// TIA Portal project "XSFW_TIA60401_A2" (V13) (continued)
VERSION : 0.1
   VAR
      x : Bool;
      x1 : Bool;
      x2 : Bool;
      x3 : Bool;
      x4 : Bool;
      x5 : Bool;
      x6 : Bool;
      x7 : Bool;
      x8 : Bool;
      x9 : Bool;
      x10 : Bool;
      x11 : Bool;
      x12 : Bool;
      x13 : Bool;
      x14 : Bool;
      x15 : Bool;
      x16 : Bool;
      x17 : Bool;
      x18 : Bool;
      x19 : Bool;
      x20 : Bool;
      x21 : Bool;
      x22 : Bool;
      x23 : Bool;
      x24 : Bool;
      x25 : Bool;
      x26 : Bool;
      x27 : Bool;
      x28 : Bool;
      x29 : Bool;
      x30 : Bool;
      x31 : Bool;
      x32 : Bool;
      x33 : Bool;
      x34 : Bool;
      x35 : Bool;
      x36 : Bool;
      x37 : Bool;
      x38 : Bool;
      x39 : Bool;
      x40 : Bool;
      x41 : Bool;
      x42 : Bool;
      x43 : Bool;
      x44 : Bool;
      x45 : Bool;
      x46 : Bool;
      x47 : Bool;
      x48 : Bool;
      x49 : Bool;
      x50 : Bool;
      x51 : Bool;
      x52 : Bool;
      x53 : Bool;
      x54 : Bool;
      x55 : Bool;
      x56 : Bool;
      x57 : Bool;
      x58 : Bool;
      x59 : Bool;
      x60 : Bool;
      x61 : Bool;
      x62 : Bool;
      x63 : Bool;
      x64 : Bool;
      x65 : Bool;
      x66 : Bool;
      x67 : Bool;
      x68 : Bool;
      x69 : Bool;
      x70 : Bool;
      x71 : Bool;
      x72 : Bool;
      x73 : Bool;
      x74 : Bool;
      x75 : Bool;
      x76 : Bool;
      x77 : Bool;
      x78 : Bool;
      x79 : Bool;
      x80 : Bool;
      x81 : Bool;
      x82 : Bool;
      x83 : Bool;
      x84 : Bool;
      x85 : Bool;
      x86 : Bool;
      x87 : Bool;
      x88 : Bool;
      x89 : Bool;
      x90 : Bool;
      x91 : Bool;
      x92 : Bool;
      x93 : Bool;
      x94 : Bool;
      x95 : Bool;
      x96 : Bool;
      x97 : Bool;
      x98 : Bool;
      x99 : Bool;
      x100 : Bool;
      x101 : Bool;
      x102 : Bool;
      x103 : Bool;
      x104 : Bool;
      x105 : Bool;
      x106 : Bool;
      x107 : Bool;
      x108 : Bool;
      x109 : Bool;
      x110 : Bool;
      x111 : Bool;
      x112 : Bool;
      x113 : Bool;
      x114 : Bool;
      x115 : Bool;
      x116 : Bool;
      x117 : Bool;
      x118 : Bool;
      x119 : Bool;
      x120 : Bool;
      x121 : Bool;
      x122 : Bool;
      x123 : Bool;
      x124 : Bool;
      x125 : Bool;
      x126 : Bool;
      x127 : Bool;
      x128 : Bool;
      x129 : Bool;
      x130 : Bool;
      x131 : Bool;
      x132 : Bool;
      x133 : Bool;
      x134 : Bool;
      x135 : Bool;
      x136 : Bool;
      x137 : Bool;
      x138 : Bool;
      x139 : Bool;
      x140 : Bool;
      x141 : Bool;
      x142 : Bool;
      x143 : Bool;
      x144 : Bool;
      x145 : Bool;
      x146 : Bool;
      x147 : Bool;
      x148 : Bool;
      x149 : Bool;
      x150 : Bool;
      x151 : Bool;
      x152 : Bool;
      x153 : Bool;
      x154 : Bool;
      x155 : Bool;
      x156 : Bool;
      x157 : Bool;
      x158 : Bool;
      x159 : Bool;
      x160 : Bool;
      x161 : Bool;
      x162 : Bool;
      x163 : Bool;
      x164 : Bool;
      x165 : Bool;
      x166 : Bool;
      x167 : Bool;
      x168 : Bool;
      x169 : Bool;
      x170 : Bool;
      x171 : Bool;
      x172 : Bool;
      x173 : Bool;
      x174 : Bool;
      x175 : Bool;
      x176 : Bool;
      x177 : Bool;
      x178 : Bool;
      x179 : Bool;
      x180 : Bool;
      x181 : Bool;
      x182 : Bool;
      x183 : Bool;
      x184 : Bool;
      x185 : Bool;
      x186 : Bool;
      x187 : Bool;
      x188 : Bool;
      x189 : Bool;
      x190 : Bool;
      x191 : Bool;
      x192 : Bool;
      x193 : Bool;
      x194 : Bool;
      x195 : Bool;
      x196 : Bool;
      x197 : Bool;
      x198 : Bool;
      x199 : Bool;
   END_VAR
BEGIN
END_DATA_BLOCK

DATA_BLOCK "DB_COM_REC_AUX"   // DB37
{ S7_Optimized_Access := 'FALSE' }
VERSION : 0.1
   VAR
      x : Bool;
      x1 : Bool;
      x2 : Bool;
      x3 : Bool;
      x4 : Bool;
      x5 : Bool;
      x6 : Bool;
      x7 : Bool;
      x8 : Bool;
      x9 : Bool;
      x10 : Bool;
      x11 : Bool;
      x12 : Bool;
      x13 : Bool;
      x14 : Bool;
      x15 : Bool;
      x16 : Bool;
      x17 : Bool;
      x18 : Bool;
      x19 : Bool;
      x20 : Bool;
      x21 : Bool;
      x22 : Bool;
      x23 : Bool;
      x24 : Bool;
      x25 : Bool;
      x26 : Bool;
      x27 : Bool;
      x28 : Bool;
      x29 : Bool;
      x30 : Bool;
      x31 : Bool;
      x32 : Bool;
      x33 : Bool;
      x34 : Bool;
      x35 : Bool;
      x36 : Bool;
      x37 : Bool;
      x38 : Bool;
      x39 : Bool;
      x40 : Bool;
      x41 : Bool;
      x42 : Bool;
      x43 : Bool;
      x44 : Bool;
      x45 : Bool;
      x46 : Bool;
      x47 : Bool;
      x48 : Bool;
      x49 : Bool;
      x50 : Bool;
      x51 : Bool;
      x52 : Bool;
      x53 : Bool;
      x54 : Bool;
      x55 : Bool;
      x56 : Bool;
      x57 : Bool;
      x58 : Bool;
      x59 : Bool;
      x60 : Bool;
      x61 : Bool;
      x62 : Bool;
      x63 : Bool;
      x64 : Bool;
      x65 : Bool;
      x66 : Bool;
      x67 : Bool;
      x68 : Bool;
      x69 : Bool;
      x70 : Bool;
      x71 : Bool;
      x72 : Bool;
      x73 : Bool;
      x74 : Bool;
      x75 : Bool;
      x76 : Bool;
      x77 : Bool;
      x78 : Bool;
      x79 : Bool;
      x80 : Bool;
      x81 : Bool;
      x82 : Bool;
      x83 : Bool;
      x84 : Bool;
      x85 : Bool;
      x86 : Bool;
      x87 : Bool;
      x88 : Bool;
      x89 : Bool;
      x90 : Bool;
      x91 : Bool;
      x92 : Bool;
      x93 : Bool;
      x94 : Bool;
      x95 : Bool;
      x96 : Bool;
      x97 : Bool;
      x98 : Bool;
      x99 : Bool;
      x100 : Bool;
      x101 : Bool;
      x102 : Bool;
      x103 : Bool;
      x104 : Bool;
      x105 : Bool;
      x106 : Bool;
      x107 : Bool;
      x108 : Bool;
      x109 : Bool;
      x110 : Bool;
      x111 : Bool;
      x112 : Bool;
      x113 : Bool;
      x114 : Bool;
      x115 : Bool;
      x116 : Bool;
      x117 : Bool;
      x118 : Bool;
      x119 : Bool;
      x120 : Bool;
      x121 : Bool;
      x122 : Bool;
      x123 : Bool;
      x124 : Bool;
      x125 : Bool;
      x126 : Bool;
      x127 : Bool;
      x128 : Bool;
      x129 : Bool;
      x130 : Bool;
      x131 : Bool;
      x132 : Bool;
      x133 : Bool;
      x134 : Bool;
      x135 : Bool;
      x136 : Bool;
      x137 : Bool;
      x138 : Bool;
      x139 : Bool;
      x140 : Bool;
      x141 : Bool;
      x142 : Bool;
      x143 : Bool;
      x144 : Bool;
      x145 : Bool;
      x146 : Bool;
      x147 : Bool;
      x148 : Bool;
      x149 : Bool;
      x150 : Bool;
      x151 : Bool;
      x152 : Bool;
      x153 : Bool;
      x154 : Bool;
      x155 : Bool;
      x156 : Bool;
      x157 : Bool;
      x158 : Bool;
      x159 : Bool;
      x160 : Bool;
      x161 : Bool;
      x162 : Bool;
      x163 : Bool;
      x164 : Bool;
      x165 : Bool;
      x166 : Bool;
      x167 : Bool;
      x168 : Bool;
      x169 : Bool;
      x170 : Bool;
      x171 : Bool;
      x172 : Bool;
      x173 : Bool;
      x174 : Bool;
      x175 : Bool;
      x176 : Bool;
      x177 : Bool;
      x178 : Bool;
      x179 : Bool;
      x180 : Bool;
      x181 : Bool;
      x182 : Bool;
      x183 : Bool;
      x184 : Bool;
      x185 : Bool;
      x186 : Bool;
      x187 : Bool;
      x188 : Bool;
      x189 : Bool;
      x190 : Bool;
      x191 : Bool;
      x192 : Bool;
      x193 : Bool;
      x194 : Bool;
      x195 : Bool;
      x196 : Bool;
      x197 : Bool;
      x198 : Bool;
      x199 : Bool;
   END_VAR
BEGIN
END_DATA_BLOCK

DATA_BLOCK "DB_BIT_VIDA"   // DB38
{ S7_Optimized_Access := 'FALSE' }
VERSION : 0.1
   VAR
      x : Bool;
      x1 : Bool;
      x2 : Bool;
      x3 : Bool;
      x4 : Bool;
      x5 : Bool;
      x6 : Bool;
      x7 : Bool;
      x8 : Bool;
      x9 : Bool;
      x10 : Bool;
      x11 : Bool;
      x12 : Bool;
      x13 : Bool;
      x14 : Bool;
      x15 : Bool;
      x16 : Bool;
      x17 : Bool;
      x18 : Bool;
      x19 : Bool;
      x20 : Bool;
      x21 : Bool;
      x22 : Bool;
      x23 : Bool;
      x24 : Bool;
      x25 : Bool;
      x26 : Bool;
      x27 : Bool;
      x28 : Bool;
      x29 : Bool;
      x30 : Bool;
      x31 : Bool;
      x32 : Bool;
      x33 : Bool;
      x34 : Bool;
      x35 : Bool;
      x36 : Bool;
      x37 : Bool;
      x38 : Bool;
      x39 : Bool;
      x40 : Bool;
      x41 : Bool;
      x42 : Bool;
      x43 : Bool;
      x44 : Bool;
      x45 : Bool;
      x46 : Bool;
      x47 : Bool;
      x48 : Bool;
      x49 : Bool;
      x50 : Bool;
      x51 : Bool;
      x52 : Bool;
      x53 : Bool;
      x54 : Bool;
      x55 : Bool;
      x56 : Bool;
      x57 : Bool;
      x58 : Bool;
      x59 : Bool;
      x60 : Bool;
      x61 : Bool;
      x62 : Bool;
      x63 : Bool;
      x64 : Bool;
      x65 : Bool;
      x66 : Bool;
      x67 : Bool;
      x68 : Bool;
      x69 : Bool;
      x70 : Bool;
      x71 : Bool;
      x72 : Bool;
      x73 : Bool;
      x74 : Bool;
      x75 : Bool;
      x76 : Bool;
      x77 : Bool;
      x78 : Bool;
      x79 : Bool;
      x80 : Bool;
      x81 : Bool;
      x82 : Bool;
      x83 : Bool;
      x84 : Bool;
      x85 : Bool;
      x86 : Bool;
      x87 : Bool;
      x88 : Bool;
      x89 : Bool;
      x90 : Bool;
      x91 : Bool;
      x92 : Bool;
      x93 : Bool;
      x94 : Bool;
      x95 : Bool;
      x96 : Bool;
      x97 : Bool;
      x98 : Bool;
      x99 : Bool;
      x100 : Bool;
      x101 : Bool;
      x102 : Bool;
      x103 : Bool;
      x104 : Bool;
      x105 : Bool;
      x106 : Bool;
      x107 : Bool;
      x108 : Bool;
      x109 : Bool;
      x110 : Bool;
      x111 : Bool;
      x112 : Bool;
      x113 : Bool;
      x114 : Bool;
      x115 : Bool;
      x116 : Bool;
      x117 : Bool;
      x118 : Bool;
      x119 : Bool;
      x120 : Bool;
      x121 : Bool;
      x122 : Bool;
      x123 : Bool;
      x124 : Bool;
      x125 : Bool;
      x126 : Bool;
      x127 : Bool;
      x128 : Bool;
      x129 : Bool;
      x130 : Bool;
      x131 : Bool;
      x132 : Bool;
      x133 : Bool;
      x134 : Bool;
      x135 : Bool;
      x136 : Bool;
      x137 : Bool;
      x138 : Bool;
      x139 : Bool;
      x140 : Bool;
      x141 : Bool;
      x142 : Bool;
      x143 : Bool;
      x144 : Bool;
      x145 : Bool;
      x146 : Bool;
      x147 : Bool;
      x148 : Bool;
      x149 : Bool;
      x150 : Bool;
      x151 : Bool;
      x152 : Bool;
      x153 : Bool;
      x154 : Bool;
      x155 : Bool;
      x156 : Bool;
      x157 : Bool;
      x158 : Bool;
      x159 : Bool;
      x160 : Bool;
      x161 : Bool;
      x162 : Bool;
      x163 : Bool;
      x164 : Bool;
      x165 : Bool;
      x166 : Bool;
      x167 : Bool;
      x168 : Bool;
      x169 : Bool;
      x170 : Bool;
      x171 : Bool;
      x172 : Bool;
      x173 : Bool;
      x174 : Bool;
      x175 : Bool;
      x176 : Bool;
      x177 : Bool;
      x178 : Bool;
      x179 : Bool;
      x180 : Bool;
      x181 : Bool;
      x182 : Bool;
      x183 : Bool;
      x184 : Bool;
      x185 : Bool;
      x186 : Bool;
      x187 : Bool;
      x188 : Bool;
      x189 : Bool;
      x190 : Bool;
      x191 : Bool;
      x192 : Bool;
      x193 : Bool;
      x194 : Bool;
      x195 : Bool;
      x196 : Bool;
      x197 : Bool;
      x198 : Bool;
      x199 : Bool;
   END_VAR
BEGIN
END_DATA_BLOCK

DATA_BLOCK "AuxiliarAlarmasMTA"   // DB47
{ S7_Optimized_Access := 'FALSE' }
VERSION : 0.1
   VAR
      AlarmaNueva : Bool;
      AlarmaPresente : Bool;
      SinAlarmas : Bool;
      Flanco_Bit_Vida : Bool;
      Falla_Comunicacion : Bool;
      Bit_Vida_Recibido : Bool;
      ReconocerTodas : Bool;
      Bit_Vida_Enviado : Bool;
   END_VAR
BEGIN
END_DATA_BLOCK

DATA_BLOCK "AlarmasDoblePantalla"   // DB86
{ S7_Optimized_Access := 'FALSE' }
VERSION : 0.1
   VAR
      x0 : Bool;
      x1 : Bool;
      x2 : Bool;
      x3 : Bool;
      x4 : Bool;
      x5 : Bool;
      x6 : Bool;
      x7 : Bool;
      r0 : Bool;
      r1 : Bool;
      r2 : Bool;
      r3 : Bool;
      r4 : Bool;
      r5 : Bool;
      r6 : Bool;
      r7 : Bool;
      x8 : Bool;
      x9 : Bool;
      x10 : Bool;
      x11 : Bool;
      x12 : Bool;
      x13 : Bool;
      x14 : Bool;
      x15 : Bool;
      r8 : Bool;
      r9 : Bool;
      r10 : Bool;
      r11 : Bool;
      r12 : Bool;
      r13 : Bool;
      r14 : Bool;
      r15 : Bool;
      x16 : Bool;
      x17 : Bool;
      x18 : Bool;
      x19 : Bool;
      x20 : Bool;
      x21 : Bool;
      x22 : Bool;
      x23 : Bool;
      r16 : Bool;
      r17 : Bool;
      r18 : Bool;
      r19 : Bool;
      r20 : Bool;
      r21 : Bool;
      r22 : Bool;
      r23 : Bool;
      x24 : Bool;
      x25 : Bool;
      x26 : Bool;
      x27 : Bool;
      x28 : Bool;
      x29 : Bool;
      x30 : Bool;
      x31 : Bool;
      r24 : Bool;
      r25 : Bool;
      r26 : Bool;
      r27 : Bool;
      r28 : Bool;
      r29 : Bool;
      r30 : Bool;
      r31 : Bool;
      x32 : Bool;
      x33 : Bool;
      x34 : Bool;
      x35 : Bool;
      x36 : Bool;
      x37 : Bool;
      x38 : Bool;
      x39 : Bool;
      r32 : Bool;
      r33 : Bool;
      r34 : Bool;
      r35 : Bool;
      r36 : Bool;
      r37 : Bool;
      r38 : Bool;
      r39 : Bool;
      x40 : Bool;
      x41 : Bool;
      x42 : Bool;
      x43 : Bool;
      x44 : Bool;
      x45 : Bool;
      x46 : Bool;
      x47 : Bool;
      r40 : Bool;
      r41 : Bool;
      r42 : Bool;
      r43 : Bool;
      r44 : Bool;
      r45 : Bool;
      r46 : Bool;
      r47 : Bool;
      x48 : Bool;
      x49 : Bool;
      x50 : Bool;
      x51 : Bool;
      x52 : Bool;
      x53 : Bool;
      x54 : Bool;
      x55 : Bool;
      r48 : Bool;
      r49 : Bool;
      r50 : Bool;
      r51 : Bool;
      r52 : Bool;
      r53 : Bool;
      r54 : Bool;
      r55 : Bool;
      x56 : Bool;
      x57 : Bool;
      x58 : Bool;
      x59 : Bool;
      x60 : Bool;
      x61 : Bool;
      x62 : Bool;
      x63 : Bool;
      r56 : Bool;
      r57 : Bool;
      r58 : Bool;
      r59 : Bool;
      r60 : Bool;
      r61 : Bool;
      r62 : Bool;
      r63 : Bool;
      x64 : Bool;
      x65 : Bool;
      x66 : Bool;
      x67 : Bool;
      x68 : Bool;
      x69 : Bool;
      x70 : Bool;
      x71 : Bool;
      r64 : Bool;
      r65 : Bool;
      r66 : Bool;
      r67 : Bool;
      r68 : Bool;
      r69 : Bool;
      r70 : Bool;
      r71 : Bool;
      x72 : Bool;
      x73 : Bool;
      x74 : Bool;
      x75 : Bool;
      x76 : Bool;
      x77 : Bool;
      x78 : Bool;
      x79 : Bool;
      r72 : Bool;
      r73 : Bool;
      r74 : Bool;
      r75 : Bool;
      r76 : Bool;
      r77 : Bool;
      r78 : Bool;
      r79 : Bool;
      x80 : Bool;
      x81 : Bool;
      x82 : Bool;
      x83 : Bool;
      x84 : Bool;
      x85 : Bool;
      x86 : Bool;
      x87 : Bool;
      r80 : Bool;
      r81 : Bool;
      r82 : Bool;
      r83 : Bool;
      r84 : Bool;
      r85 : Bool;
      r86 : Bool;
      r87 : Bool;
      x88 : Bool;
      x89 : Bool;
      x90 : Bool;
      x91 : Bool;
      x92 : Bool;
      x93 : Bool;
      x94 : Bool;
      x95 : Bool;
      r88 : Bool;
      r89 : Bool;
      r90 : Bool;
      r91 : Bool;
      r92 : Bool;
      r93 : Bool;
      r94 : Bool;
      r95 : Bool;
      x96 : Bool;
      x97 : Bool;
      x98 : Bool;
      x99 : Bool;
      x100 : Bool;
      x101 : Bool;
      x102 : Bool;
      x103 : Bool;
      r96 : Bool;
      r97 : Bool;
      r98 : Bool;
      r99 : Bool;
      r100 : Bool;
      r101 : Bool;
      r102 : Bool;
      r103 : Bool;
      x104 : Bool;
      x105 : Bool;
      x106 : Bool;
      x107 : Bool;
      x108 : Bool;
      x109 : Bool;
      x110 : Bool;
      x111 : Bool;
      r104 : Bool;
      r105 : Bool;
      r106 : Bool;
      r107 : Bool;
      r108 : Bool;
      r109 : Bool;
      r110 : Bool;
      r111 : Bool;
      x112 : Bool;
      x113 : Bool;
      x114 : Bool;
      x115 : Bool;
      x116 : Bool;
      x117 : Bool;
      x118 : Bool;
      x119 : Bool;
      r112 : Bool;
      r113 : Bool;
      r114 : Bool;
      r115 : Bool;
      r116 : Bool;
      r117 : Bool;
      r118 : Bool;
      r119 : Bool;
      x120 : Bool;
      x121 : Bool;
      x122 : Bool;
      x123 : Bool;
      x124 : Bool;
      x125 : Bool;
      x126 : Bool;
      x127 : Bool;
      r120 : Bool;
      r121 : Bool;
      r122 : Bool;
      r123 : Bool;
      r124 : Bool;
      r125 : Bool;
      r126 : Bool;
      r127 : Bool;
      x128 : Bool;
      x129 : Bool;
      x130 : Bool;
      x131 : Bool;
      x132 : Bool;
      x133 : Bool;
      x134 : Bool;
      x135 : Bool;
      r128 : Bool;
      r129 : Bool;
      r130 : Bool;
      r131 : Bool;
      r132 : Bool;
      r133 : Bool;
      r134 : Bool;
      r135 : Bool;
      x136 : Bool;
      x137 : Bool;
      x138 : Bool;
      x139 : Bool;
      x140 : Bool;
      x141 : Bool;
      x142 : Bool;
      x143 : Bool;
      r136 : Bool;
      r137 : Bool;
      r138 : Bool;
      r139 : Bool;
      r140 : Bool;
      r141 : Bool;
      r142 : Bool;
      r143 : Bool;
      x144 : Bool;
      x145 : Bool;
      x146 : Bool;
      x147 : Bool;
      x148 : Bool;
      x149 : Bool;
      x150 : Bool;
      x151 : Bool;
      r144 : Bool;
      r145 : Bool;
      r146 : Bool;
      r147 : Bool;
      r148 : Bool;
      r149 : Bool;
      r150 : Bool;
      r151 : Bool;
      x152 : Bool;
      x153 : Bool;
      x154 : Bool;
      x155 : Bool;
      x156 : Bool;
      x157 : Bool;
      x158 : Bool;
      x159 : Bool;
      r152 : Bool;
      r153 : Bool;
      r154 : Bool;
      r155 : Bool;
      r156 : Bool;
      r157 : Bool;
      r158 : Bool;
      r159 : Bool;
      x160 : Bool;
      x161 : Bool;
      x162 : Bool;
      x163 : Bool;
      x164 : Bool;
      x165 : Bool;
      x166 : Bool;
      x167 : Bool;
      r160 : Bool;
      r161 : Bool;
      r162 : Bool;
      r163 : Bool;
      r164 : Bool;
      r165 : Bool;
      r166 : Bool;
      r167 : Bool;
      x168 : Bool;
      x169 : Bool;
      x170 : Bool;
      x171 : Bool;
      x172 : Bool;
      x173 : Bool;
      x174 : Bool;
      x175 : Bool;
      r168 : Bool;
      r169 : Bool;
      r170 : Bool;
      r171 : Bool;
      r172 : Bool;
      r173 : Bool;
      r174 : Bool;
      r175 : Bool;
      x176 : Bool;
      x177 : Bool;
      x178 : Bool;
      x179 : Bool;
      x180 : Bool;
      x181 : Bool;
      x182 : Bool;
      x183 : Bool;
      r176 : Bool;
      r177 : Bool;
      r178 : Bool;
      r179 : Bool;
      r180 : Bool;
      r181 : Bool;
      r182 : Bool;
      r183 : Bool;
      x184 : Bool;
      x185 : Bool;
      x186 : Bool;
      x187 : Bool;
      x188 : Bool;
      x189 : Bool;
      x190 : Bool;
      x191 : Bool;
      r184 : Bool;
      r185 : Bool;
      r186 : Bool;
      r187 : Bool;
      r188 : Bool;
      r189 : Bool;
      r190 : Bool;
      r191 : Bool;
      x192 : Bool;
      x193 : Bool;
      x194 : Bool;
      x195 : Bool;
      x196 : Bool;
      x197 : Bool;
      x198 : Bool;
      x199 : Bool;
      r192 : Bool;
      r193 : Bool;
      r194 : Bool;
      r195 : Bool;
      r196 : Bool;
      r197 : Bool;
      r198 : Bool;
      r199 : Bool;
   END_VAR
BEGIN
END_DATA_BLOCK

DATA_BLOCK "CFGSirena"   // DB91
{ S7_Optimized_Access := 'FALSE' }
VERSION : 0.1
   VAR
      Motivo1 : Bool;
      Motivo2 : Bool;
      Motivo3 : Bool;
      Motivo4 : Bool;
      Motivo5 : Bool;
      Motivo6 : Bool;
      Motivo7 : Bool;
      Motivo8 : Bool;
      Motivo9 : Bool;
      Motivo10 : Bool;
      Motivo11 : Bool;
      Motivo12 : Bool;
      Motivo13 : Bool;
      Motivo14 : Bool;
      Motivo15 : Bool;
      Motivo16 : Bool;
      Motivo17 : Bool;
      Motivo18 : Bool;
      Motivo19 : Bool;
      Motivo20 : Bool;
      Motivo21 : Bool;
      Motivo22 : Bool;
      Motivo23 : Bool;
      Motivo24 : Bool;
   END_VAR
BEGIN
END_DATA_BLOCK

// folder: Bloques Estándar/Boosters

DATA_BLOCK "Boosters Gral"   // DB62
{ S7_Optimized_Access := 'FALSE' }
VERSION : 0.1
   VAR
      SegBoost1 : Int;
      SegBoost2 : Int;
      MinBoost1 : Int;
      MinBoost2 : Int;
      HorasBoost1 : DInt;
      HorasBoost2 : DInt;
      HorasLim : DInt;
      TiempoAyudaON_PANEL : Word;
      TiempoAyudaOFF_PANEL : Word;
      TiempoAyudaON : S5Time;
      TiempoAyudaOFF : S5Time;
      LimArrPrio2 : Real;
      LimArrPrio1 : Real;
      LimParPrio2 : Real;
      LimParPrio1 : Real;
      Ctrl_Analogico : Bool;
   END_VAR
BEGIN
END_DATA_BLOCK

// folder: Compresores/Alta

DATA_BLOCK "AuxiliarVLV"   // DB10
{ S7_Optimized_Access := 'FALSE' }
VERSION : 0.1
   VAR
      DejarAbrirVLV1 : Bool;
      DejarAbrirVLV2 : Bool;
      DejarAbrirVLV3 : Bool;
      DejarAbrirVLV4 : Bool;
      DejarAbrirVLV5 : Bool;
      DejarAbrirVLV6 : Bool;
   END_VAR
BEGIN
END_DATA_BLOCK

DATA_BLOCK "DB-PurgaComAlta"   // DB53
{ S7_Optimized_Access := 'FALSE' }
VERSION : 0.1
   VAR
      Habil_PurgaBellis : Bool;
      Habil_PurgaABC2 : Bool;
      Habil_PurgaABC3 : Bool;
      Habil_PurgaABC4 : Bool;
      Habil_PurgaABC5 : Bool;
      Habil_PurgaABC1 : Bool;
      Toff_PurgaBellis : Word;
      Ton_PurgaBellis : Word;
      Toff_PurgaABC2 : Word;
      Ton_PurgaABC2 : Word;
      Toff_PurgaABC3 : Word;
      Ton_PurgaABC3 : Word;
      Toff_PurgaABC4 : Word;
      Ton_PurgaABC4 : Word;
      Toff_PurgaABC5 : Word;
      Ton_PurgaABC5 : Word;
      Toff_PurgaABC1 : Word;
      Ton_PurgaABC1 : Word;
      Prueba_PurgaBellis : Bool;
      Prueba_PurgaABC2 : Bool;
      Prueba_PurgaABC3 : Bool;
      Prueba_PurgaABC4 : Bool;
      Prueba_PurgaABC5 : Bool;
      Prueba_PurgaABC1 : Bool;
   END_VAR
BEGIN
END_DATA_BLOCK

DATA_BLOCK "Agregado Bellis"   // DB63
{ S7_Optimized_Access := 'FALSE' }
VERSION : 0.1
   VAR
      ExcesoTiempo : S5Time;
      ForzarCompleta : Bool;
      QuitarForzado : Bool;
      ExcesoTiempoPanel : Int;
   END_VAR
BEGIN
END_DATA_BLOCK

DATA_BLOCK "PanelCompALTA MTA"   // DB75
{ S7_Optimized_Access := 'FALSE' }
VERSION : 0.1
   VAR
      DB_VAR : Int;
   END_VAR
BEGIN
END_DATA_BLOCK

DATA_BLOCK "DB-CompAltaDatos"   // DB88
{ S7_Optimized_Access := 'FALSE' }
VERSION : 0.1
   VAR
      Req : Int;
      F_Osc_1seg : Bool;
      MinParGen : Int;
      PanMchCmp1 : Bool;
      PanMchCmp2 : Bool;
      PanMchCmp3 : Bool;
      PanMchCmp4 : Bool;
      PanMchCmp5 : Bool;
      PanMchCmp6 : Bool;
      TON_ParGen : Bool;
      TON_ParGen_Lim : Bool;
      ValorParGen : Int;
      Aut1 : Bool;
      Aut2 : Bool;
      Aut3 : Bool;
      Aut4 : Bool;
      Aut5 : Bool;
      Aut6 : Bool;
      TON_ParGenMem : Bool;
      CgaPrsCrt : Bool;
   END_VAR
BEGIN
END_DATA_BLOCK

DATA_BLOCK "FallasCmpALTA"   // DB89
{ S7_Optimized_Access := 'FALSE' }
VERSION : 0.1
   VAR
      FaGen1 : Bool;
      FaGen2 : Bool;
      FaGen3 : Bool;
      FaGen4 : Bool;
      FaGen5 : Bool;
      FaGen6 : Bool;
      FaGen : Bool;
   END_VAR
BEGIN
END_DATA_BLOCK

DATA_BLOCK "CompALTA-MTA"   // DB121
{ S7_Optimized_Access := 'FALSE' }
VERSION : 0.1
   VAR
      FallaGral : Bool;
      FallaCompresor1 : Bool;
      FallaCompresor2 : Bool;
      FallaCompresor3 : Bool;
      FallaCompresor4 : Bool;
      FallaCompresor5 : Bool;
      FallaCompresor6 : Bool;
      EncenderAutoComp1 : Bool;
      EncenderAutoComp2 : Bool;
      EncenderAutoComp3 : Bool;
      EncenderAutoComp4 : Bool;
      EncenderAutoComp5 : Bool;
      EncenderAutoComp6 : Bool;
      IndVCmp1 : Bool;
      IndVCmp2 : Bool;
      IndVCmp3 : Bool;
      IndVCmp4 : Bool;
      IndVCmp5 : Bool;
      IndVCmp6 : Bool;
      IndRCmp1 : Bool;
      IndRCmp2 : Bool;
      IndRCmp3 : Bool;
      IndRCmp4 : Bool;
      IndRCmp5 : Bool;
      IndRCmp6 : Bool;
      CmpReq : Word;
      IndMarchaCmp1 : Bool;
      IndMarchaCmp2 : Bool;
      IndMarchaCmp3 : Bool;
      IndMarchaCmp4 : Bool;
      IndMarchaCmp5 : Bool;
      IndMarchaCmp6 : Bool;
      OvrLimP1 : Bool;
      OvrLimP2 : Bool;
      OvrLimP3 : Bool;
      OvrLimP4 : Bool;
      OvrLimP5 : Bool;
      OvrLimP6 : Bool;
      UndLimP1 : Bool;
      RESETPrioridades : Bool;
      UndLimP2 : Bool;
      UndLimP3 : Bool;
      UndLimP4 : Bool;
      UndLimP5 : Bool;
      UndLimP6 : Bool;
      PrsMed : Real;
      MchP1 : Bool;
      MchP2 : Bool;
      MchP3 : Bool;
      MchP4 : Bool;
      MchP5 : Bool;
      MchP6 : Bool;
      CgaP1 : Bool;
      CgaP2 : Bool;
      CgaP3 : Bool;
      CgaP4 : Bool;
      CgaP5 : Bool;
      CgaP6 : Bool;
      VRealCmp1 : Int;
      Reserva : Int;
      VRealCmp2 : Int;
      Reserva1 : Int;
      VRealCmp3 : Int;
      Reserva2 : Int;
      VRealCmp4 : Int;
      Reserva3 : Int;
      VRealCmp5 : Int;
      Reserva4 : Int;
      VRealCmp6 : Int;
      Reserva5 : Int;
      ReqMch1 : Bool;
      ReqMch2 : Bool;
      ReqMch3 : Bool;
      ReqMch4 : Bool;
      ReqMch5 : Bool;
      ReqMch6 : Bool;
      SinReq1 : Bool;
      SinReq2 : Bool;
      SinReq3 : Bool;
      SinReq4 : Bool;
      SinReq5 : Bool;
      SinReq6 : Bool;
      ManP1 : Bool;
      ManP2 : Bool;
      ManP3 : Bool;
      ManP4 : Bool;
      ManP5 : Bool;
      ManP6 : Bool;
      CicloIni : Bool;
      ReqCga1 : Bool;
      ReqCga2 : Bool;
      ReqCga3 : Bool;
      ReqCga4 : Bool;
      ReqCga5 : Bool;
      ReqCga6 : Bool;
      ReqCrr : Int;
      AnimCMP1 : Int;
      AnimCMP2 : Int;
      AnimCMP3 : Int;
      AnimCMP4 : Int;
      AnimCMP5 : Int;
      AnimCMP6 : Int;
      AnimGen : Int;
      Reset : Bool;
      UltPriDis : Int;
      CntReqIte : Int;
      CntReqCrr : Int;
      CntCmpDisp : Int;
      IndVP1 : Bool;
      IndVP2 : Bool;
      IndVP3 : Bool;
      IndVP4 : Bool;
      IndVP5 : Bool;
      IndVP6 : Bool;
      OvrLimPCRT : Bool;
      UndLimPCRT : Bool;
   END_VAR
BEGIN
END_DATA_BLOCK

DATA_BLOCK "DBParamCmpALTA-MTA"   // DB122
{ S7_Optimized_Access := 'FALSE' }
VERSION : 0.1
   VAR
      LimSupP1 : Real;
      LimSupP2 : Real;
      LimSupP3 : Real;
      LimSupP4 : Real;
      LimSupP5 : Real;
      LimSupP6 : Real;
      LimInfP1 : Real;
      LimInfP2 : Real;
      LimInfP3 : Real;
      LimInfP4 : Real;
      LimInfP5 : Real;
      LimInfP6 : Real;
      DelPrs : Real;
      HstPrs : Real;
      PrsMax : Real;
      HstPrsCrt : Real;
      LimSupPCRT : Real;
      LimInfPCRT : Real;
      LMedia1 : Real;
      LMedia2 : Real;
      LMedia3 : Real;
      LMedia4 : Real;
      LMedia5 : Real;
      LMedia6 : Real;
      MediaHist : Real;
      TempCritEnclav : Real;
   END_VAR
BEGIN
END_DATA_BLOCK

DATA_BLOCK "DBTiemposCmpAltaMTA"   // DB123
{ S7_Optimized_Access := 'FALSE' }
VERSION : 0.1
   VAR
      FNueReqIni : Bool;
      Reserva2 : Bool;
      Reserva3 : Bool;
      Reserva4 : Bool;
      Reserva5 : Bool;
      TVAC : S5Time;
      TVACPANEL : Int;
      TVACPEsc : Int;
      RetSinRec : S5Time;
      RetSinRecPANEL : Int;
      RetSinRecPEsc : Int;
   END_VAR
BEGIN
END_DATA_BLOCK

DATA_BLOCK "Sopladoras"   // DB124
{ S7_Optimized_Access := 'FALSE' }
VERSION : 0.1
   VAR
      Sop1 : Bool;
      Sop2 : Bool;
      Sop3 : Bool;
      TStopSop : S5Time;
      TStopSopPanel : Int;
      NinSOP : Bool;
      ReqSp1 : Int;
      ReqSp2 : Int;
      ReqSp3 : Int;
      ReqIni : Int;
      FinClcReq : Bool;
   END_VAR
BEGIN
END_DATA_BLOCK

DATA_BLOCK "DB-PrioridadesCmpAlta"   // DB125
{ S7_Optimized_Access := 'FALSE' }
VERSION : 0.1
   VAR
      Vcmp0 : Int;
      Vcmp1 : Int;
      Vcmp2 : Int;
      Vcmp3 : Int;
      Vcmp4 : Int;
      Vcmp5 : Int;
      Vcmp6 : Int;
      fDecPri1 : Bool;
      fDecPri2 : Bool;
      fDecPri3 : Bool;
      fDecPri4 : Bool;
      fDecPri5 : Bool;
      fDecPri6 : Bool;
      fIncPri1 : Bool;
      fIncPri2 : Bool;
      fIncPri3 : Bool;
      fIncPri4 : Bool;
      fIncPri5 : Bool;
      fIncPri6 : Bool;
      IncPri1 : Bool;
      IncPri2 : Bool;
      IncPri3 : Bool;
      IncPri4 : Bool;
      IncPri5 : Bool;
      IncPri6 : Bool;
      DecPri1 : Bool;
      DecPri2 : Bool;
      DecPri3 : Bool;
      DecPri4 : Bool;
      DecPri5 : Bool;
      DecPri6 : Bool;
   END_VAR
BEGIN
END_DATA_BLOCK

DATA_BLOCK "DB-AccionamientosCmpAlta"   // DB126
{ S7_Optimized_Access := 'FALSE' }
VERSION : 0.1
   VAR
      DB_VAR : Int;
   END_VAR
BEGIN
END_DATA_BLOCK

DATA_BLOCK "PanelCmpAlta"   // DB135
{ S7_Optimized_Access := 'FALSE' }
VERSION : 0.1
   VAR
      AnimMenu1 : Int;
      AnimMenu2 : Int;
      AnimMenu3 : Int;
      AnimMenu4 : Int;
      AnimMenu5 : Int;
      AnimMenu6 : Int;
      SPON1 : Real;
      SPON2 : Real;
      SPON3 : Real;
      SPON4 : Real;
      SPON5 : Real;
      SPON6 : Real;
      SPOFF1 : Real;
      SPOFF2 : Real;
      SPOFF3 : Real;
      SPOFF4 : Real;
      SPOFF5 : Real;
      SPOFF6 : Real;
      MantMC001 : Bool;
      MantMC002 : Bool;
      MantMC003 : Bool;
      MantMC004 : Bool;
      MantMC005 : Bool;
      MantMC006 : Bool;
      MachaMC001 : Bool;
      MachaMC002 : Bool;
      MachaMC003 : Bool;
      MachaMC004 : Bool;
      MachaMC005 : Bool;
      MachaMC006 : Bool;
      MarchaPanelMC001 : Bool;
      MarchaPanelMC002 : Bool;
      MarchaPanelMC003 : Bool;
      MarchaPanelMC004 : Bool;
      MarchaPanelMC005 : Bool;
      MarchaPanelMC006 : Bool;
      ParadaPanelMC001 : Bool;
      ParadaPanelMC002 : Bool;
      ParadaPanelMC003 : Bool;
      ParadaPanelMC004 : Bool;
      ParadaPanelMC005 : Bool;
      ParadaPanelMC006 : Bool;
      MediaCargaBellis : Bool;
      AbrirVLV1 : Bool;
      AbrirVLV2 : Bool;
      AbrirVLV3 : Bool;
      AbrirVLV4 : Bool;
      AbrirVLV5 : Bool;
      AbrirVLV6 : Bool;
      AbrirVLV3b : Bool;
   END_VAR
BEGIN
END_DATA_BLOCK

DATA_BLOCK "ModoManualCompAlta"   // DB136
{ S7_Optimized_Access := 'FALSE' }
VERSION : 0.1
   VAR
      MarchaFPanel1 : Bool;
      MarchaFPanel2 : Bool;
      MarchaFPanel3 : Bool;
      MarchaFPanel4 : Bool;
      MarchaFPanel5 : Bool;
      MarchaFPanel6 : Bool;
      ParadaFPanel1 : Bool;
      ParadaFPanel2 : Bool;
      ParadaFPanel3 : Bool;
      ParadaFPanel4 : Bool;
      ParadaFPanel5 : Bool;
      ParadaFPanel6 : Bool;
      OrdenMarchaForzada1 : Bool;
      OrdenMarchaForzada2 : Bool;
      OrdenMarchaForzada3 : Bool;
      OrdenMarchaForzada4 : Bool;
      OrdenMarchaForzada5 : Bool;
      OrdenMarchaForzada6 : Bool;
      VlvManual1 : Bool;
      VlvManual2 : Bool;
      VlvManual3 : Bool;
      VlvManual4 : Bool;
      VlvManual5 : Bool;
      VlvManual6 : Bool;
      SPON1 : Real;
      SPON2 : Real;
      SPON3 : Real;
      SPON4 : Real;
      SPON5 : Real;
      SPON6 : Real;
      SPOFF1 : Real;
      SPOFF2 : Real;
      SPOFF3 : Real;
      SPOFF4 : Real;
      SPOFF5 : Real;
      SPOFF6 : Real;
      SPON3b : Real;
      SPOFF3b : Real;
      VlvManual3b : Bool;
   END_VAR
BEGIN
END_DATA_BLOCK

// folder: Compresores/Alta/Máquina de Estados

DATA_BLOCK "EstadosCmpALTA-MTA"   // DB120
{ S7_Optimized_Access := 'FALSE' }
VERSION : 0.1
   VAR
      _1s1 : Bool;
      _1s2 : Bool;
      _1s3 : Bool;
      _1s4 : Bool;
      _1s5 : Bool;
      _1s6 : Bool;
      _1s7 : Bool;
      _1s8 : Bool;
      _1s9 : Bool;
      _1s10 : Bool;
      _1sReserva2 : Bool;
      _1sReserva3 : Bool;
      _1sReserva4 : Bool;
      _1sReserva5 : Bool;
      _1sReserva6 : Bool;
      _1sReserva7 : Bool;
      _2s1 : Bool;
      _2s2 : Bool;
      _2s3 : Bool;
      _2s4 : Bool;
      _2s5 : Bool;
      _2s6 : Bool;
      _2s7 : Bool;
      _2s8 : Bool;
      _2s9 : Bool;
      _2s10 : Bool;
      _2sReserva2 : Bool;
      _2sReserva3 : Bool;
      _2sReserva4 : Bool;
      _2sReserva5 : Bool;
      _2sReserva6 : Bool;
      _2sReserva7 : Bool;
      _3s1 : Bool;
      _3s2 : Bool;
      _3s3 : Bool;
      _3s4 : Bool;
      _3s5 : Bool;
      _3s6 : Bool;
      _3s7 : Bool;
      _3s8 : Bool;
      _3s9 : Bool;
      _3s10 : Bool;
      _3Reserva2 : Bool;
      _3Reserva3 : Bool;
      _3Reserva4 : Bool;
      _3Reserva5 : Bool;
      _3Reserva6 : Bool;
      _3Reserva7 : Bool;
      _4s1 : Bool;
      _4s2 : Bool;
      _4s3 : Bool;
      _4s4 : Bool;
      _4s5 : Bool;
      _4s6 : Bool;
      _4s7 : Bool;
      _4s8 : Bool;
      _4s9 : Bool;
      _4s10 : Bool;
      _4sReserva2 : Bool;
      _4sReserva3 : Bool;
      _4sReserva4 : Bool;
      _4sReserva5 : Bool;
      _4sReserva6 : Bool;
      _4sReserva7 : Bool;
      _5s1 : Bool;
      _5s2 : Bool;
      _5s3 : Bool;
      _5s4 : Bool;
      _5s5 : Bool;
      _5s6 : Bool;
      _5s7 : Bool;
      _5s8 : Bool;
      _5s9 : Bool;
      _5s10 : Bool;
      _5sReserva2 : Bool;
      _5sReserva3 : Bool;
      _5sReserva4 : Bool;
      _5sReserva5 : Bool;
      _5sReserva6 : Bool;
      _5sReserva7 : Bool;
      _6s1 : Bool;
      _6s2 : Bool;
      _6s3 : Bool;
      _6s4 : Bool;
      _6s5 : Bool;
      _6s6 : Bool;
      _6s7 : Bool;
      _6s8 : Bool;
      _6s9 : Bool;
      _6s10 : Bool;
      _6sReserva2 : Bool;
      _6sReserva3 : Bool;
      _6sReserva4 : Bool;
      _6sReserva5 : Bool;
      _6sReserva6 : Bool;
      _6sReserva7 : Bool;
      _0s1 : Bool;
      _0s2 : Bool;
      _0s3 : Bool;
      _0s4 : Bool;
      _0s5 : Bool;
      _0s6 : Bool;
      _0s7 : Bool;
      _0s8 : Bool;
      _0s9 : Bool;
      _0s10 : Bool;
      _0sReserva2 : Bool;
      _0sReserva3 : Bool;
      _0sReserva4 : Bool;
      _0sReserva5 : Bool;
      _0sReserva6 : Bool;
      _0sReserva7 : Bool;
   END_VAR
BEGIN
END_DATA_BLOCK

DATA_BLOCK "Concatenadoras"   // DB127
{ S7_Optimized_Access := 'FALSE' }
VERSION : 0.1
   VAR
      _1c1 : Bool;
      _1c2 : Bool;
      _1c3 : Bool;
      _1c4 : Bool;
      _1c5 : Bool;
      _1c6 : Bool;
      _1c7 : Bool;
      _1c8 : Bool;
      _1c9 : Bool;
      _1c10 : Bool;
      _1cReserva2 : Bool;
      _1cReserva3 : Bool;
      _1cReserva4 : Bool;
      _1cReserva5 : Bool;
      _1cReserva6 : Bool;
      _1cReserva7 : Bool;
      _2c1 : Bool;
      _2c2 : Bool;
      _2c3 : Bool;
      _2c4 : Bool;
      _2c5 : Bool;
      _2c6 : Bool;
      _2c7 : Bool;
      _2c8 : Bool;
      _2c9 : Bool;
      _2c10 : Bool;
      _2cReserva2 : Bool;
      _2cReserva3 : Bool;
      _2cReserva4 : Bool;
      _2cReserva5 : Bool;
      _2cReserva6 : Bool;
      _2cReserva7 : Bool;
      _3c1 : Bool;
      _3c2 : Bool;
      _3c3 : Bool;
      _3c4 : Bool;
      _3c5 : Bool;
      _3c6 : Bool;
      _3c7 : Bool;
      _3c8 : Bool;
      _3c9 : Bool;
      _3c10 : Bool;
      _3cReserva2 : Bool;
      _3cReserva3 : Bool;
      _3cReserva4 : Bool;
      _3cReserva5 : Bool;
      _3cReserva6 : Bool;
      _3cReserva7 : Bool;
      _4c1 : Bool;
      _4c2 : Bool;
      _4c3 : Bool;
      _4c4 : Bool;
      _4c5 : Bool;
      _4c6 : Bool;
      _4c7 : Bool;
      _4c8 : Bool;
      _4c9 : Bool;
      _4c10 : Bool;
      _4cReserva2 : Bool;
      _4cReserva3 : Bool;
      _4cReserva4 : Bool;
      _4cReserva5 : Bool;
      _4cReserva6 : Bool;
      _4cReserva7 : Bool;
      _5c1 : Bool;
      _5c2 : Bool;
      _5c3 : Bool;
      _5c4 : Bool;
      _5c5 : Bool;
      _5c6 : Bool;
      _5c7 : Bool;
      _5c8 : Bool;
      _5c9 : Bool;
      _5c10 : Bool;
      _5cReserva2 : Bool;
      _5cReserva3 : Bool;
      _5cReserva4 : Bool;
      _5cReserva5 : Bool;
      _5cReserva6 : Bool;
      _5cReserva7 : Bool;
      _6c1 : Bool;
      _6c2 : Bool;
      _6c3 : Bool;
      _6c4 : Bool;
      _6c5 : Bool;
      _6c6 : Bool;
      _6c7 : Bool;
      _6c8 : Bool;
      _6c9 : Bool;
      _6c10 : Bool;
      _6cReserva2 : Bool;
      _6cReserva3 : Bool;
      _6cReserva4 : Bool;
      _6cReserva5 : Bool;
      _6cReserva6 : Bool;
      _6cReserva7 : Bool;
      _0c1 : Bool;
      _0c2 : Bool;
      _0c3 : Bool;
      _0c4 : Bool;
      _0c5 : Bool;
      _0c6 : Bool;
      _0c7 : Bool;
      _0c8 : Bool;
      _0c9 : Bool;
      _0c10 : Bool;
      _0cReserva2 : Bool;
      _0cReserva3 : Bool;
      _0cReserva4 : Bool;
      _0cReserva5 : Bool;
      _0cReserva6 : Bool;
      _0cReserva7 : Bool;
   END_VAR
BEGIN
END_DATA_BLOCK

